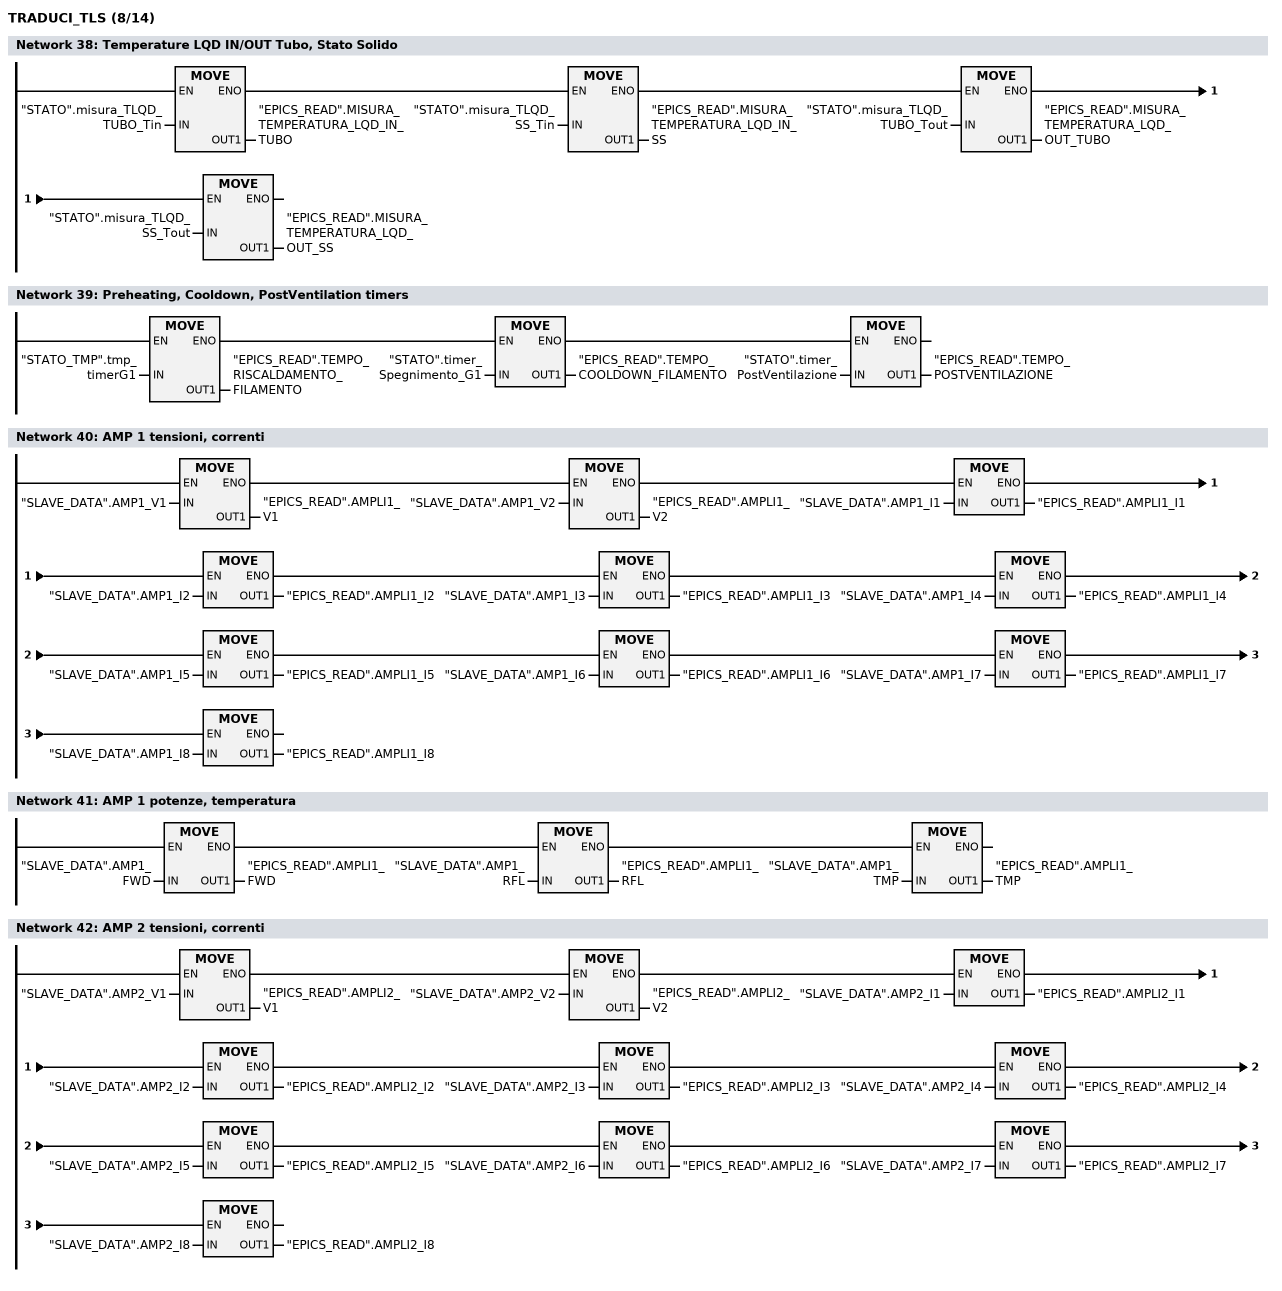
   RUNG wire#powerrail
      Move(in := "STATO".misura_TLQD_TUBO_Tin, out1 => "EPICS_READ".MISURA_TEMPERATURA_LQD_IN_TUBO)
      Move(in := "STATO".misura_TLQD_SS_Tin, out1 => "EPICS_READ".MISURA_TEMPERATURA_LQD_IN_SS)
      Move(in := "STATO".misura_TLQD_TUBO_Tout, out1 => "EPICS_READ".MISURA_TEMPERATURA_LQD_OUT_TUBO)
      Move(in := "STATO".misura_TLQD_SS_Tout, out1 => "EPICS_READ".MISURA_TEMPERATURA_LQD_OUT_SS)
   END_RUNG
   // the same network as SCL:
   "EPICS_READ".MISURA_TEMPERATURA_LQD_IN_TUBO := "STATO".misura_TLQD_TUBO_Tin;
   "EPICS_READ".MISURA_TEMPERATURA_LQD_IN_SS := "STATO".misura_TLQD_SS_Tin;
   "EPICS_READ".MISURA_TEMPERATURA_LQD_OUT_TUBO := "STATO".misura_TLQD_TUBO_Tout;
   "EPICS_READ".MISURA_TEMPERATURA_LQD_OUT_SS := "STATO".misura_TLQD_SS_Tout;
END_REGION

REGION Network 39: Preheating, Cooldown, PostVentilation timers
   RUNG wire#powerrail
      Move(in := "STATO_TMP".tmp_timerG1, out1 => "EPICS_READ".TEMPO_RISCALDAMENTO_FILAMENTO)
      Move(in := "STATO".timer_Spegnimento_G1, out1 => "EPICS_READ".TEMPO_COOLDOWN_FILAMENTO)
      Move(in := "STATO".timer_PostVentilazione, out1 => "EPICS_READ".TEMPO_POSTVENTILAZIONE)
   END_RUNG
   // the same network as SCL:
   "EPICS_READ".TEMPO_RISCALDAMENTO_FILAMENTO := "STATO_TMP".tmp_timerG1;
   "EPICS_READ".TEMPO_COOLDOWN_FILAMENTO := "STATO".timer_Spegnimento_G1;
   "EPICS_READ".TEMPO_POSTVENTILAZIONE := "STATO".timer_PostVentilazione;
END_REGION

REGION Network 40: AMP 1 tensioni, correnti
   RUNG wire#powerrail
      Move(in := "SLAVE_DATA".AMP1_V1, out1 => "EPICS_READ".AMPLI1_V1)
      Move(in := "SLAVE_DATA".AMP1_V2, out1 => "EPICS_READ".AMPLI1_V2)
      Move(in := "SLAVE_DATA".AMP1_I1, out1 => "EPICS_READ".AMPLI1_I1)
      Move(in := "SLAVE_DATA".AMP1_I2, out1 => "EPICS_READ".AMPLI1_I2)
      Move(in := "SLAVE_DATA".AMP1_I3, out1 => "EPICS_READ".AMPLI1_I3)
      Move(in := "SLAVE_DATA".AMP1_I4, out1 => "EPICS_READ".AMPLI1_I4)
      Move(in := "SLAVE_DATA".AMP1_I5, out1 => "EPICS_READ".AMPLI1_I5)
      Move(in := "SLAVE_DATA".AMP1_I6, out1 => "EPICS_READ".AMPLI1_I6)
      Move(in := "SLAVE_DATA".AMP1_I7, out1 => "EPICS_READ".AMPLI1_I7)
      Move(in := "SLAVE_DATA".AMP1_I8, out1 => "EPICS_READ".AMPLI1_I8)
   END_RUNG
   // the same network as SCL:
   "EPICS_READ".AMPLI1_V1 := "SLAVE_DATA".AMP1_V1;
   "EPICS_READ".AMPLI1_V2 := "SLAVE_DATA".AMP1_V2;
   "EPICS_READ".AMPLI1_I1 := "SLAVE_DATA".AMP1_I1;
   "EPICS_READ".AMPLI1_I2 := "SLAVE_DATA".AMP1_I2;
   "EPICS_READ".AMPLI1_I3 := "SLAVE_DATA".AMP1_I3;
   "EPICS_READ".AMPLI1_I4 := "SLAVE_DATA".AMP1_I4;
   "EPICS_READ".AMPLI1_I5 := "SLAVE_DATA".AMP1_I5;
   "EPICS_READ".AMPLI1_I6 := "SLAVE_DATA".AMP1_I6;
   "EPICS_READ".AMPLI1_I7 := "SLAVE_DATA".AMP1_I7;
   "EPICS_READ".AMPLI1_I8 := "SLAVE_DATA".AMP1_I8;
END_REGION

REGION Network 41: AMP 1 potenze, temperatura
   RUNG wire#powerrail
      Move(in := "SLAVE_DATA".AMP1_FWD, out1 => "EPICS_READ".AMPLI1_FWD)
      Move(in := "SLAVE_DATA".AMP1_RFL, out1 => "EPICS_READ".AMPLI1_RFL)
      Move(in := "SLAVE_DATA".AMP1_TMP, out1 => "EPICS_READ".AMPLI1_TMP)
   END_RUNG
   // the same network as SCL:
   "EPICS_READ".AMPLI1_FWD := "SLAVE_DATA".AMP1_FWD;
   "EPICS_READ".AMPLI1_RFL := "SLAVE_DATA".AMP1_RFL;
   "EPICS_READ".AMPLI1_TMP := "SLAVE_DATA".AMP1_TMP;
END_REGION

REGION Network 42: AMP 2 tensioni, correnti
   RUNG wire#powerrail
      Move(in := "SLAVE_DATA".AMP2_V1, out1 => "EPICS_READ".AMPLI2_V1)
      Move(in := "SLAVE_DATA".AMP2_V2, out1 => "EPICS_READ".AMPLI2_V2)
      Move(in := "SLAVE_DATA".AMP2_I1, out1 => "EPICS_READ".AMPLI2_I1)
      Move(in := "SLAVE_DATA".AMP2_I2, out1 => "EPICS_READ".AMPLI2_I2)
      Move(in := "SLAVE_DATA".AMP2_I3, out1 => "EPICS_READ".AMPLI2_I3)
      Move(in := "SLAVE_DATA".AMP2_I4, out1 => "EPICS_READ".AMPLI2_I4)
      Move(in := "SLAVE_DATA".AMP2_I5, out1 => "EPICS_READ".AMPLI2_I5)
      Move(in := "SLAVE_DATA".AMP2_I6, out1 => "EPICS_READ".AMPLI2_I6)
      Move(in := "SLAVE_DATA".AMP2_I7, out1 => "EPICS_READ".AMPLI2_I7)
      Move(in := "SLAVE_DATA".AMP2_I8, out1 => "EPICS_READ".AMPLI2_I8)
   END_RUNG
   // the same network as SCL:
   "EPICS_READ".AMPLI2_V1 := "SLAVE_DATA".AMP2_V1;
   "EPICS_READ".AMPLI2_V2 := "SLAVE_DATA".AMP2_V2;
   "EPICS_READ".AMPLI2_I1 := "SLAVE_DATA".AMP2_I1;
   "EPICS_READ".AMPLI2_I2 := "SLAVE_DATA".AMP2_I2;
   "EPICS_READ".AMPLI2_I3 := "SLAVE_DATA".AMP2_I3;
   "EPICS_READ".AMPLI2_I4 := "SLAVE_DATA".AMP2_I4;
   "EPICS_READ".AMPLI2_I5 := "SLAVE_DATA".AMP2_I5;
   "EPICS_READ".AMPLI2_I6 := "SLAVE_DATA".AMP2_I6;
   "EPICS_READ".AMPLI2_I7 := "SLAVE_DATA".AMP2_I7;
   "EPICS_READ".AMPLI2_I8 := "SLAVE_DATA".AMP2_I8;
END_REGION

REGION Network 43: AMP 2 potenze, temperatura
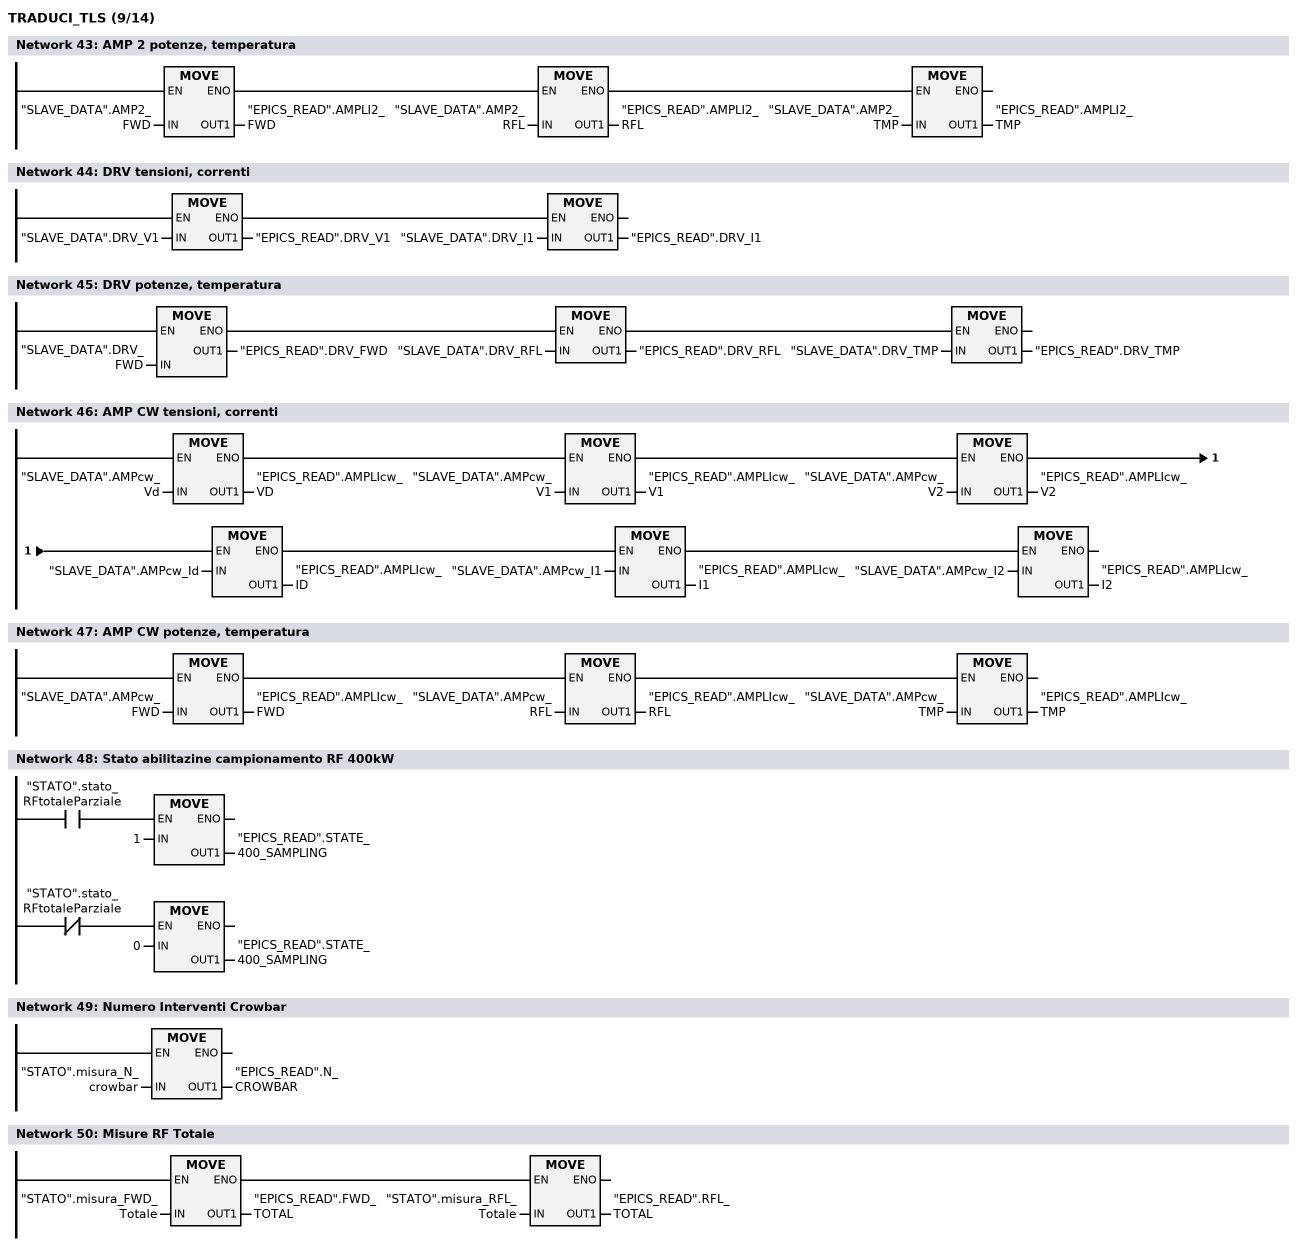
   RUNG wire#powerrail
      Move(in := "SLAVE_DATA".AMP2_FWD, out1 => "EPICS_READ".AMPLI2_FWD)
      Move(in := "SLAVE_DATA".AMP2_RFL, out1 => "EPICS_READ".AMPLI2_RFL)
      Move(in := "SLAVE_DATA".AMP2_TMP, out1 => "EPICS_READ".AMPLI2_TMP)
   END_RUNG
   // the same network as SCL:
   "EPICS_READ".AMPLI2_FWD := "SLAVE_DATA".AMP2_FWD;
   "EPICS_READ".AMPLI2_RFL := "SLAVE_DATA".AMP2_RFL;
   "EPICS_READ".AMPLI2_TMP := "SLAVE_DATA".AMP2_TMP;
END_REGION

REGION Network 44: DRV tensioni, correnti
   RUNG wire#powerrail
      Move(in := "SLAVE_DATA".DRV_V1, out1 => "EPICS_READ".DRV_V1)
      Move(in := "SLAVE_DATA".DRV_I1, out1 => "EPICS_READ".DRV_I1)
   END_RUNG
   // the same network as SCL:
   "EPICS_READ".DRV_V1 := "SLAVE_DATA".DRV_V1;
   "EPICS_READ".DRV_I1 := "SLAVE_DATA".DRV_I1;
END_REGION

REGION Network 45: DRV potenze, temperatura
   RUNG wire#powerrail
      Move(in := "SLAVE_DATA".DRV_FWD, out1 => "EPICS_READ".DRV_FWD)
      Move(in := "SLAVE_DATA".DRV_RFL, out1 => "EPICS_READ".DRV_RFL)
      Move(in := "SLAVE_DATA".DRV_TMP, out1 => "EPICS_READ".DRV_TMP)
   END_RUNG
   // the same network as SCL:
   "EPICS_READ".DRV_FWD := "SLAVE_DATA".DRV_FWD;
   "EPICS_READ".DRV_RFL := "SLAVE_DATA".DRV_RFL;
   "EPICS_READ".DRV_TMP := "SLAVE_DATA".DRV_TMP;
END_REGION

REGION Network 46: AMP CW tensioni, correnti
   RUNG wire#powerrail
      Move(in := "SLAVE_DATA".AMPcw_Vd, out1 => "EPICS_READ".AMPLIcw_VD)
      Move(in := "SLAVE_DATA".AMPcw_V1, out1 => "EPICS_READ".AMPLIcw_V1)
      Move(in := "SLAVE_DATA".AMPcw_V2, out1 => "EPICS_READ".AMPLIcw_V2)
      Move(in := "SLAVE_DATA".AMPcw_Id, out1 => "EPICS_READ".AMPLIcw_ID)
      Move(in := "SLAVE_DATA".AMPcw_I1, out1 => "EPICS_READ".AMPLIcw_I1)
      Move(in := "SLAVE_DATA".AMPcw_I2, out1 => "EPICS_READ".AMPLIcw_I2)
   END_RUNG
   // the same network as SCL:
   "EPICS_READ".AMPLIcw_VD := "SLAVE_DATA".AMPcw_Vd;
   "EPICS_READ".AMPLIcw_V1 := "SLAVE_DATA".AMPcw_V1;
   "EPICS_READ".AMPLIcw_V2 := "SLAVE_DATA".AMPcw_V2;
   "EPICS_READ".AMPLIcw_ID := "SLAVE_DATA".AMPcw_Id;
   "EPICS_READ".AMPLIcw_I1 := "SLAVE_DATA".AMPcw_I1;
   "EPICS_READ".AMPLIcw_I2 := "SLAVE_DATA".AMPcw_I2;
END_REGION

REGION Network 47: AMP CW potenze, temperatura
   RUNG wire#powerrail
      Move(in := "SLAVE_DATA".AMPcw_FWD, out1 => "EPICS_READ".AMPLIcw_FWD)
      Move(in := "SLAVE_DATA".AMPcw_RFL, out1 => "EPICS_READ".AMPLIcw_RFL)
      Move(in := "SLAVE_DATA".AMPcw_TMP, out1 => "EPICS_READ".AMPLIcw_TMP)
   END_RUNG
   // the same network as SCL:
   "EPICS_READ".AMPLIcw_FWD := "SLAVE_DATA".AMPcw_FWD;
   "EPICS_READ".AMPLIcw_RFL := "SLAVE_DATA".AMPcw_RFL;
   "EPICS_READ".AMPLIcw_TMP := "SLAVE_DATA".AMPcw_TMP;
END_REGION

REGION Network 48: Stato abilitazine campionamento RF 400kW
   RUNG wire#powerrail
      Contact( "STATO".stato_RFtotaleParziale )
      Move(in := 1, out1 => "EPICS_READ".STATE_400_SAMPLING)
   END_RUNG
   RUNG wire#powerrail
      I_Contact( "STATO".stato_RFtotaleParziale )
      Move(in := 0, out1 => "EPICS_READ".STATE_400_SAMPLING)
   END_RUNG
   // the same network as SCL:
   IF "STATO".stato_RFtotaleParziale THEN "EPICS_READ".STATE_400_SAMPLING := 1; END_IF;
   IF NOT "STATO".stato_RFtotaleParziale THEN "EPICS_READ".STATE_400_SAMPLING := 0; END_IF;
END_REGION

REGION Network 49: Numero Interventi Crowbar
   RUNG wire#powerrail
      Move(in := "STATO".misura_N_crowbar, out1 => "EPICS_READ".N_CROWBAR)
   END_RUNG
   // the same network as SCL:
   "EPICS_READ".N_CROWBAR := "STATO".misura_N_crowbar;
END_REGION

REGION Network 50: Misure RF Totale
   RUNG wire#powerrail
      Move(in := "STATO".misura_FWD_Totale, out1 => "EPICS_READ".FWD_TOTAL)
      Move(in := "STATO".misura_RFL_Totale, out1 => "EPICS_READ".RFL_TOTAL)
   END_RUNG
   // the same network as SCL:
   "EPICS_READ".FWD_TOTAL := "STATO".misura_FWD_Totale;
   "EPICS_READ".RFL_TOTAL := "STATO".misura_RFL_Totale;
END_REGION

REGION Network 51: Presenza allarme Personal Security
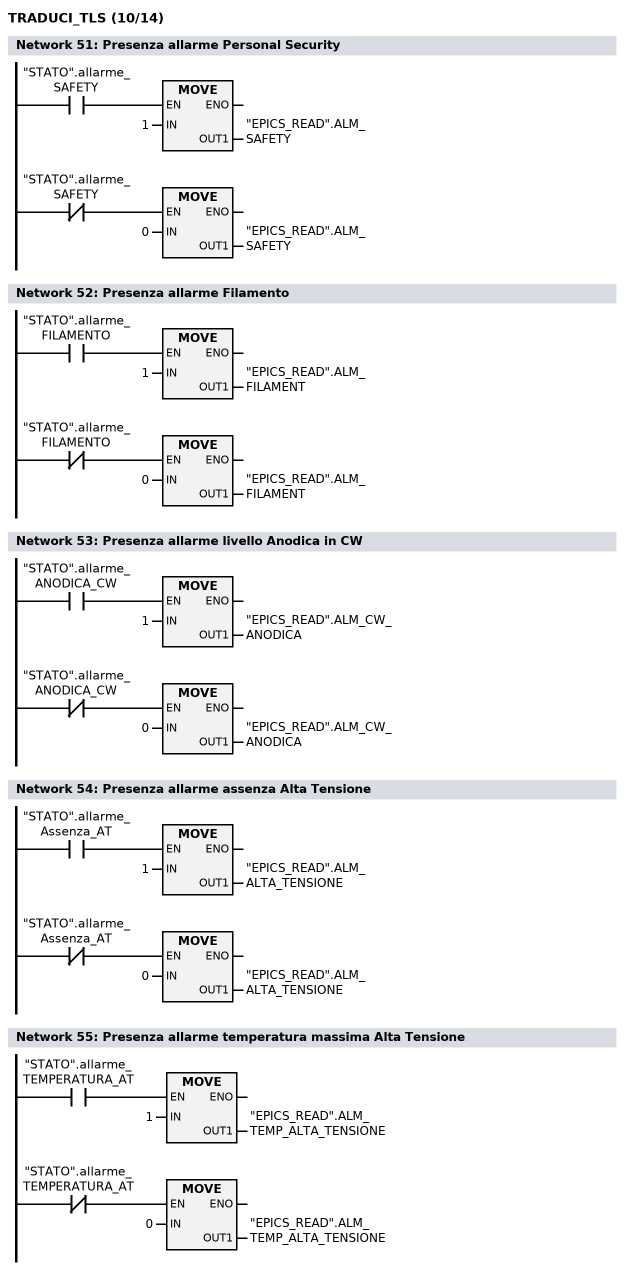
   RUNG wire#powerrail
      Contact( "STATO".allarme_SAFETY )
      Move(in := 1, out1 => "EPICS_READ".ALM_SAFETY)
   END_RUNG
   RUNG wire#powerrail
      I_Contact( "STATO".allarme_SAFETY )
      Move(in := 0, out1 => "EPICS_READ".ALM_SAFETY)
   END_RUNG
   // the same network as SCL:
   IF "STATO".allarme_SAFETY THEN "EPICS_READ".ALM_SAFETY := 1; END_IF;
   IF NOT "STATO".allarme_SAFETY THEN "EPICS_READ".ALM_SAFETY := 0; END_IF;
END_REGION

REGION Network 52: Presenza allarme Filamento
   RUNG wire#powerrail
      Contact( "STATO".allarme_FILAMENTO )
      Move(in := 1, out1 => "EPICS_READ".ALM_FILAMENT)
   END_RUNG
   RUNG wire#powerrail
      I_Contact( "STATO".allarme_FILAMENTO )
      Move(in := 0, out1 => "EPICS_READ".ALM_FILAMENT)
   END_RUNG
   // the same network as SCL:
   IF "STATO".allarme_FILAMENTO THEN "EPICS_READ".ALM_FILAMENT := 1; END_IF;
   IF NOT "STATO".allarme_FILAMENTO THEN "EPICS_READ".ALM_FILAMENT := 0; END_IF;
END_REGION

REGION Network 53: Presenza allarme livello Anodica in CW
   RUNG wire#powerrail
      Contact( "STATO".allarme_ANODICA_CW )
      Move(in := 1, out1 => "EPICS_READ".ALM_CW_ANODICA)
   END_RUNG
   RUNG wire#powerrail
      I_Contact( "STATO".allarme_ANODICA_CW )
      Move(in := 0, out1 => "EPICS_READ".ALM_CW_ANODICA)
   END_RUNG
   // the same network as SCL:
   IF "STATO".allarme_ANODICA_CW THEN "EPICS_READ".ALM_CW_ANODICA := 1; END_IF;
   IF NOT "STATO".allarme_ANODICA_CW THEN "EPICS_READ".ALM_CW_ANODICA := 0; END_IF;
END_REGION

REGION Network 54: Presenza allarme assenza Alta Tensione
   RUNG wire#powerrail
      Contact( "STATO".allarme_Assenza_AT )
      Move(in := 1, out1 => "EPICS_READ".ALM_ALTA_TENSIONE)
   END_RUNG
   RUNG wire#powerrail
      I_Contact( "STATO".allarme_Assenza_AT )
      Move(in := 0, out1 => "EPICS_READ".ALM_ALTA_TENSIONE)
   END_RUNG
   // the same network as SCL:
   IF "STATO".allarme_Assenza_AT THEN "EPICS_READ".ALM_ALTA_TENSIONE := 1; END_IF;
   IF NOT "STATO".allarme_Assenza_AT THEN "EPICS_READ".ALM_ALTA_TENSIONE := 0; END_IF;
END_REGION

REGION Network 55: Presenza allarme temperatura massima Alta Tensione
   RUNG wire#powerrail
      Contact( "STATO".allarme_TEMPERATURA_AT )
      Move(in := 1, out1 => "EPICS_READ".ALM_TEMP_ALTA_TENSIONE)
   END_RUNG
   RUNG wire#powerrail
      I_Contact( "STATO".allarme_TEMPERATURA_AT )
      Move(in := 0, out1 => "EPICS_READ".ALM_TEMP_ALTA_TENSIONE)
   END_RUNG
   // the same network as SCL:
   IF "STATO".allarme_TEMPERATURA_AT THEN "EPICS_READ".ALM_TEMP_ALTA_TENSIONE := 1; END_IF;
   IF NOT "STATO".allarme_TEMPERATURA_AT THEN "EPICS_READ".ALM_TEMP_ALTA_TENSIONE := 0; END_IF;
END_REGION

REGION Network 56: Presenza allarme Conducimetro
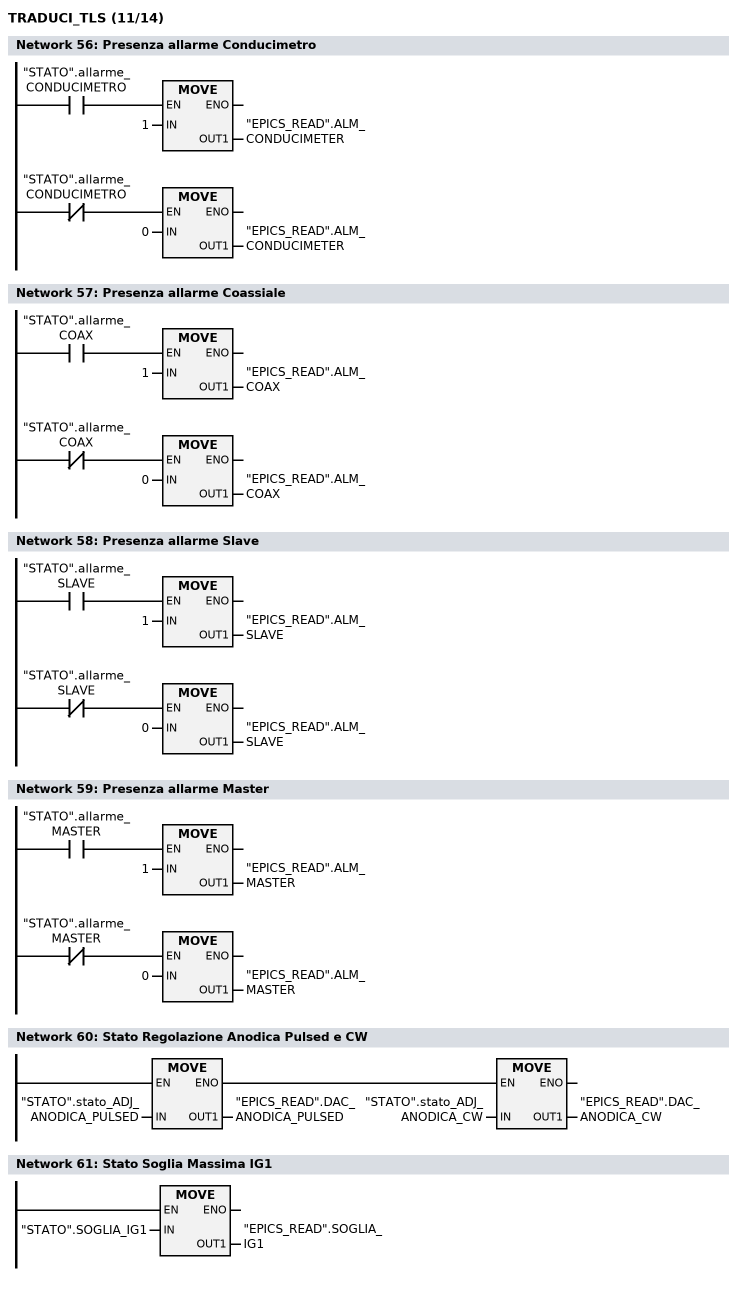
   RUNG wire#powerrail
      Contact( "STATO".allarme_CONDUCIMETRO )
      Move(in := 1, out1 => "EPICS_READ".ALM_CONDUCIMETER)
   END_RUNG
   RUNG wire#powerrail
      I_Contact( "STATO".allarme_CONDUCIMETRO )
      Move(in := 0, out1 => "EPICS_READ".ALM_CONDUCIMETER)
   END_RUNG
   // the same network as SCL:
   IF "STATO".allarme_CONDUCIMETRO THEN "EPICS_READ".ALM_CONDUCIMETER := 1; END_IF;
   IF NOT "STATO".allarme_CONDUCIMETRO THEN "EPICS_READ".ALM_CONDUCIMETER := 0; END_IF;
END_REGION

REGION Network 57: Presenza allarme Coassiale
   RUNG wire#powerrail
      Contact( "STATO".allarme_COAX )
      Move(in := 1, out1 => "EPICS_READ".ALM_COAX)
   END_RUNG
   RUNG wire#powerrail
      I_Contact( "STATO".allarme_COAX )
      Move(in := 0, out1 => "EPICS_READ".ALM_COAX)
   END_RUNG
   // the same network as SCL:
   IF "STATO".allarme_COAX THEN "EPICS_READ".ALM_COAX := 1; END_IF;
   IF NOT "STATO".allarme_COAX THEN "EPICS_READ".ALM_COAX := 0; END_IF;
END_REGION

REGION Network 58: Presenza allarme Slave
   RUNG wire#powerrail
      Contact( "STATO".allarme_SLAVE )
      Move(in := 1, out1 => "EPICS_READ".ALM_SLAVE)
   END_RUNG
   RUNG wire#powerrail
      I_Contact( "STATO".allarme_SLAVE )
      Move(in := 0, out1 => "EPICS_READ".ALM_SLAVE)
   END_RUNG
   // the same network as SCL:
   IF "STATO".allarme_SLAVE THEN "EPICS_READ".ALM_SLAVE := 1; END_IF;
   IF NOT "STATO".allarme_SLAVE THEN "EPICS_READ".ALM_SLAVE := 0; END_IF;
END_REGION

REGION Network 59: Presenza allarme Master
   RUNG wire#powerrail
      Contact( "STATO".allarme_MASTER )
      Move(in := 1, out1 => "EPICS_READ".ALM_MASTER)
   END_RUNG
   RUNG wire#powerrail
      I_Contact( "STATO".allarme_MASTER )
      Move(in := 0, out1 => "EPICS_READ".ALM_MASTER)
   END_RUNG
   // the same network as SCL:
   IF "STATO".allarme_MASTER THEN "EPICS_READ".ALM_MASTER := 1; END_IF;
   IF NOT "STATO".allarme_MASTER THEN "EPICS_READ".ALM_MASTER := 0; END_IF;
END_REGION

REGION Network 60: Stato Regolazione Anodica Pulsed e CW
   RUNG wire#powerrail
      Move(in := "STATO".stato_ADJ_ANODICA_PULSED, out1 => "EPICS_READ".DAC_ANODICA_PULSED)
      Move(in := "STATO".stato_ADJ_ANODICA_CW, out1 => "EPICS_READ".DAC_ANODICA_CW)
   END_RUNG
   // the same network as SCL:
   "EPICS_READ".DAC_ANODICA_PULSED := "STATO".stato_ADJ_ANODICA_PULSED;
   "EPICS_READ".DAC_ANODICA_CW := "STATO".stato_ADJ_ANODICA_CW;
END_REGION

REGION Network 61: Stato Soglia Massima IG1
   RUNG wire#powerrail
      Move(in := "STATO".SOGLIA_IG1, out1 => "EPICS_READ".SOGLIA_IG1)
   END_RUNG
   // the same network as SCL:
   "EPICS_READ".SOGLIA_IG1 := "STATO".SOGLIA_IG1;
END_REGION

REGION Network 62: Stato Soglia Massima IG2